               "LPMLV30_CMD_START":
                 IF NOT #statStatesInCurrentMode.resetting AND NOT #statStatesInCurrentMode.idle THEN
                   #StateChangeInProcess := TRUE;
                   #StateRequested := "LPMLV30_STATE_EXECUTE";
                   // Check if valid state for command is in use by current mode
                   IF #statStatesInCurrentMode.starting THEN
                     #statStateInternal := "LPMLV30_STATE_STARTING";
                   ELSE
                     #statStateInternal := "LPMLV30_STATE_EXECUTE";
                   END_IF;
                 ELSE
                   #diagnostics.buffer[#tempDiagnosticsBufferIndexCmd].message := #MSG_CMD_NOT_ALLOWED;
                 END_IF;
               ELSE
                 IF #diagnostics.buffer[#tempDiagnosticsBufferIndexCmd].message = #MSG_NO_MESSAGE THEN // ELSE: Message was already written in head part of message handling
                   #diagnostics.buffer[#tempDiagnosticsBufferIndexCmd].message := #MSG_CMD_NOT_ALLOWED;
                 END_IF;
             END_CASE;
           END_IF;

         "LPMLV30_STATE_UNDEFINED":
           #StateChangeInProcess := FALSE;
           #StateRequested    := "LPMLV30_STATE_STOPPED";
           #statStateInternal := "LPMLV30_STATE_STOPPED";
         ELSE
           ; // Undefined state
       END_CASE;
     END_IF; // End: state machine

     //-------------------------------------------------
     // Message handling for state manager: foot part
     //-------------------------------------------------
     IF #statStateInternal <> #statStateCurrentOld THEN // ELSE: States were not changed
       IF #tempDiagnosticsBufferIndexCmd >= 0 AND #tempDiagnosticsBufferIndexCmd <= "LPMLV30_DIAG_BUFFER_UPPER_LIM" THEN
         IF #diagnostics.buffer[#tempDiagnosticsBufferIndexCmd].message = #MSG_NO_MESSAGE THEN
           #diagnostics.buffer[#tempDiagnosticsBufferIndexCmd].message := #MSG_STATE_CHANGED_SUCCESSFULLY;
         END_IF;
       END_IF;
       IF #tempDiagnosticsBufferIndexSC >= 0 AND #tempDiagnosticsBufferIndexSC <= "LPMLV30_DIAG_BUFFER_UPPER_LIM" THEN
         IF #diagnostics.buffer[#tempDiagnosticsBufferIndexSC].message = #MSG_NO_MESSAGE THEN
           #diagnostics.buffer[#tempDiagnosticsBufferIndexSC].message := #MSG_STATE_CHANGED_SUCCESSFULLY;
         END_IF;
       END_IF;
     END_IF; // End: message handling for state manager: foot part
   END_IF; // End: As from second cycle
   // End: State manager

   //--------------------------------------------------------------------------------------------------
   // Write outputs including boolean interface outputs 
   //--------------------------------------------------------------------------------------------------
   IF #statUnitModeCurrentInternal <> #statUnitModeCurrentInternalOld THEN // Check if new unit mode is selected
     #ProductionModeActive  := FALSE;
     #MaintenanceModeActive := FALSE;
     #ManualModeActive      := FALSE;
     #UserMode01Active      := FALSE;
     #UserMode02Active      := FALSE;
     #UserMode03Active      := FALSE;
     #UserMode04Active      := FALSE;
     #UserMode05Active      := FALSE;
     #UserMode06Active      := FALSE;
     #UserMode07Active      := FALSE;
     #UserMode08Active      := FALSE;
     // #UserMode09Active := FALSE;
     // #UserMode10Active := FALSE;
     // #UserMode11Active := FALSE;
     // #UserMode13Active := FALSE;
     // #UserMode14Active := FALSE;
     // #UserMode15Active := FALSE;
     // #UserMode16Active := FALSE;
     // #UserMode17Active := FALSE;
     // #UserMode18Active := FALSE;
     // #UserMode19Active := FALSE;
     // #UserMode20Active := FALSE;
     // #UserMode21Active := FALSE;
     // #UserMode22Active := FALSE;
     // #UserMode23Active := FALSE;
     // #UserMode24Active := FALSE;
     // #UserMode25Active := FALSE;
     // #UserMode26Active := FALSE;
     // #UserMode27Active := FALSE;
     // #UserMode28Active := FALSE;

     CASE #statUnitModeCurrentInternal OF // Set new bit for current unit mode
       "LPMLV30_MODE_PRODUCTION":
         #ProductionModeActive := TRUE;
       "LPMLV30_MODE_MAINTENANCE":
         #MaintenanceModeActive := TRUE;
       "LPMLV30_MODE_MANUAL":
         #ManualModeActive := TRUE;
       "LPMLV30_MODE_USER_01":
         #UserMode01Active := TRUE;
       "LPMLV30_MODE_USER_02":
         #UserMode02Active := TRUE;
       "LPMLV30_MODE_USER_03":
         #UserMode03Active := TRUE;
       "LPMLV30_MODE_USER_04":
         #UserMode04Active := TRUE;
       "LPMLV30_MODE_USER_05":
         #UserMode05Active := TRUE;
       "LPMLV30_MODE_USER_06":
         #UserMode06Active := TRUE;
       "LPMLV30_MODE_USER_07":
         #UserMode07Active := TRUE;
       "LPMLV30_MODE_USER_08":
         #UserMode08Active := TRUE;
       // LPMLV30_MODE_USER_09:
       //   #UserMode09Active := TRUE;
       // LPMLV30_MODE_USER_10:
       //   #UserMode10Active := TRUE;
       // LPMLV30_MODE_USER_11:
       //   #UserMode11Active := TRUE;
       // LPMLV30_MODE_USER_12:
       //   #UserMode12Active := TRUE;
       // LPMLV30_MODE_USER_13:
       //   #UserMode13Active := TRUE;
       // LPMLV30_MODE_USER_14:
       //   #UserMode14Active := TRUE;
       // LPMLV30_MODE_USER_15:
       //   #UserMode15Active := TRUE;
       // LPMLV30_MODE_USER_16:
       //   #UserMode16Active := TRUE;
       // LPMLV30_MODE_USER_17:
       //   #UserMode17Active := TRUE;
       // LPMLV30_MODE_USER_18:
       //   #UserMode18Active := TRUE;
       // LPMLV30_MODE_USER_19:
       //   #UserMode19Active := TRUE;
       // LPMLV30_MODE_USER_20:
       //   #UserMode20Active := TRUE;
       // LPMLV30_MODE_USER_21:
       //   #UserMode21Active := TRUE;
       // LPMLV30_MODE_USER_22:
       //   #UserMode22Active := TRUE;
       // LPMLV30_MODE_USER_23:
       //   #UserMode23Active := TRUE;
       // LPMLV30_MODE_USER_24:
       //   #UserMode25Active := TRUE;
       // LPMLV30_MODE_USER_25:
       //   #UserMode25Active := TRUE;
       // LPMLV30_MODE_USER_26:
       //   #UserMode26Active := TRUE;
       // LPMLV30_MODE_USER_27:
       //   #UserMode27Active := TRUE;
       // LPMLV30_MODE_USER_28:
       //   #UserMode28Active := TRUE;
       ELSE
         ; // No bit is set
     END_CASE;

     #statUnitModeCurrentInternalOld := #statUnitModeCurrentInternal;
   END_IF;

   IF #statStateInternal <> #statStateInternalOld THEN // Check if new state is selected 
     #StateCurrent := #statStateInternal; // Set output

     // Set states of boolean interface out
     // Delete old state  
     #ClearingStateActive     := FALSE;
     #StoppedStateActive      := FALSE;
     #StartingStateActive     := FALSE;
     #IdleStateActive         := FALSE;
     #SuspendedStateActive    := FALSE;
     #ExecuteStateActive      := FALSE;
     #StoppingStateActive     := FALSE;
     #AbortingStateActive     := FALSE;
     #AbortedStateActive      := FALSE;
     #HoldingStateActive      := FALSE;
     #HeldStateActive         := FALSE;
     #UnholdingStateActive    := FALSE;
     #SuspendingStateActive   := FALSE;
     #UnsuspendingStateActive := FALSE;
     #ResettingStateActive    := FALSE;
     #CompletingStateActive   := FALSE;
     #CompleteStateActive     := FALSE;

     // Set new state
     CASE #statStateInternal OF
       "LPMLV30_STATE_CLEARING":
         #ClearingStateActive := TRUE;
       "LPMLV30_STATE_STOPPED":
         #StoppedStateActive := TRUE;
       "LPMLV30_STATE_STARTING":
         #StartingStateActive := TRUE;
       "LPMLV30_STATE_IDLE":
         #IdleStateActive := TRUE;
       "LPMLV30_STATE_SUSPENDED":
         #SuspendedStateActive := TRUE;
       "LPMLV30_STATE_EXECUTE":
         #ExecuteStateActive := TRUE;
       "LPMLV30_STATE_STOPPING":
         #StoppingStateActive := TRUE;
       "LPMLV30_STATE_ABORTING":
         #AbortingStateActive := TRUE;
       "LPMLV30_STATE_ABORTED":
         #AbortedStateActive := TRUE;
       "LPMLV30_STATE_HOLDING":
         #HoldingStateActive := TRUE;
       "LPMLV30_STATE_HELD":
         #HeldStateActive := TRUE;
       "LPMLV30_STATE_UNHOLDING":
         #UnholdingStateActive := TRUE;
       "LPMLV30_STATE_SUSPENDING":
         #SuspendingStateActive := TRUE;
       "LPMLV30_STATE_UNSUSPENDING":
         #UnsuspendingStateActive := TRUE;
       "LPMLV30_STATE_RESETTING":
         #ResettingStateActive := TRUE;
       "LPMLV30_STATE_COMPLETING":
         #CompletingStateActive := TRUE;
       "LPMLV30_STATE_COMPLETE":
         #CompleteStateActive := TRUE;
       ELSE
         ;
     END_CASE; // End: Set new state

     #statStateInternalOld := #statStateInternal;
   END_IF;// End: Write boolean interface outputs

   #diagnostics.bufferIndex := #tempDiagnosticsBufferIndex; // Temporary variable is used during block execution -> Copy back/Set output
   IF #statFirstCycle THEN
     #statFirstCycle := FALSE;
   END_IF;

   // Save values for edge detection
   IF #statUnitModeChangeRequest THEN
     #statUnitModeOld := #statUnitMode;
   END_IF;
   IF #statCmdChangeRequest THEN
     #statCntrlCmdOld := #tempCntrlCmd;
   END_IF;
   IF #statStateInternal <> #statStateCurrentOld THEN
     #statStateCurrentOld := #statStateInternal;
   END_IF;

   //============================================================================================================
   // End of function block: LPMLV30_UnitModeStateManager
   //============================================================================================================
END_FUNCTION_BLOCK

FUNCTION_BLOCK "LPMLV30_UnitModeStateTimes"   // FB30101, SCL
TITLE = LPMLV30_UnitModeStateTimes
{ S7_Optimized_Access := 'TRUE' }
AUTHOR : APC_ERLF
FAMILY : OMAC
// Support: tech.team.motioncontrol@siemens.com 
// Fax: +49 (0) 9131/98-1297
   VAR_INPUT
      UnitModeCurrent : DInt := 0;   // Current unit mode
      StateCurrent : DInt := 0;   // Current state
      resetTimes : Bool := false;   // State change from FALSE to TRUE (rising edge) resets unit mode/state times and cumulative times
   END_VAR
   VAR_OUTPUT
      ModeCurrentTime : Array[0.."LPMLV30_MODES_UPPER_LIM"] of DInt;   // Current time for all modes in seconds
      ModeCumulativeTime : Array[0.."LPMLV30_MODES_UPPER_LIM"] of DInt;   // Cumulative time for all modes in seconds
      StateCurrentTime : Array[0.."LPMLV30_MODES_UPPER_LIM", 0.."LPMLV30_STATES_UPPER_LIM"] of DInt;   // Current time for all states in seconds
      StateCumulativeTime : Array[0.."LPMLV30_MODES_UPPER_LIM", 0.."LPMLV30_STATES_UPPER_LIM"] of DInt;   // Cumulative time for all states in seconds
      actualTimeCurrentMode : DInt;   // Actual time for current mode in seconds
      cumulativeTimeCurrentMode : DInt;   // Cumulative time for current mode in seconds
      actualTimeCurrentStates : Array[0.."LPMLV30_STATES_UPPER_LIM"] of DInt;   // Actual time for all states in current mode in seconds
      cumulativeTimeCurrentStates : Array[0.."LPMLV30_STATES_UPPER_LIM"] of DInt;   // Cumulative time for all states in current mode in seconds
      AccTimeSinceReset : DInt;   // Accumulated time since last reset in seconds
   END_VAR
   VAR
      statUnitModeCurrentOld : DInt := 0;   // For edge detection
      statStateCurrentOld : DInt := 0;   // For edge detection
      statResetTimesOld : Bool := false;   // For edge detection
      statStartingPointMeasureRuntime : LReal := 0.0;   // Saved value of runtime system function
      statRuntime : LReal := 0.0;   // Runtime variable
      statFirstCycle : Bool := true;   // First cycle of run
   END_VAR
   VAR_TEMP
      tempI : Int;   // Loop counter
      tempJ : Int;   // Loop counter
      tempMeasuredRuntime : LReal;   // Return value of RUNTIME instruction
      tempRuntimeIntegerPart : DInt;   // Runtime variable (integer part)
      tempUnitModeCurrent : DInt;   // Verified input value
      tempStateCurrent : DInt;   // Verified input value
   END_VAR
BEGIN
   //============================================================================================================
   // SIEMENS AG
   // (c)Copyright 2015 All Rights Reserved
   //------------------------------------------------------------------------------------------------------------
   // Library: LPMLV30
   // Tested with: S7-1200 with FW version V4.1, S7-1500 with FW version V1.7
   // Engineering: TIA Portal V13 SP1
   // Restrictions: ---
   // Requirements: S7-1200 / S7-1500
   // Functionality: Determination of unit modes and states times (current and also cumulative times)
   //------------------------------------------------------------------------------------------------------------
   // Change log table:
   // Version  Date        Expert in charge    Changes applied
   // 03.00.01 29.05.2015  RK                  First released version 
   //============================================================================================================
   // Function block: LPMLV30_UnitModeStateTimes
   //============================================================================================================

   IF #statFirstCycle OR (#resetTimes AND NOT #statResetTimesOld) THEN
     // Reset times structures
     FOR #tempI := "LPMLV30_MODE_INVALID" TO "LPMLV30_MODES_UPPER_LIM" DO
       #ModeCurrentTime[#tempI] := 0;
       IF NOT #statFirstCycle THEN // Do only with rising edge at resetTimes
         #ModeCumulativeTime[#tempI] := 0;
       END_IF;
       FOR #tempJ := "LPMLV30_STATE_UNDEFINED" TO "LPMLV30_STATES_UPPER_LIM" DO
         #StateCurrentTime[#tempI, #tempJ] := 0;
         IF NOT #statFirstCycle THEN // Do only with rising edge at resetTimes
           #StateCumulativeTime[#tempI, #tempJ] := 0;
         END_IF;
       END_FOR;
     END_FOR;
     IF NOT #statFirstCycle THEN // Do only with rising edge at resetTimes
       #AccTimeSinceReset := 0;
     END_IF;

     // Reset additional outputs
     #actualTimeCurrentMode := 0;
     IF NOT #statFirstCycle THEN // Do only with rising edge at resetTimes
       #cumulativeTimeCurrentMode := 0;
     END_IF;
     FOR #tempI := "LPMLV30_STATE_UNDEFINED" TO "LPMLV30_STATES_UPPER_LIM" DO
       #actualTimeCurrentStates[#tempI] := 0;
       IF NOT #statFirstCycle THEN // Do only with rising edge at resetTimes
         #cumulativeTimeCurrentStates[#tempI] := 0;
       END_IF;
     END_FOR;

     // Set starting point for calculation of elapsed seconds
     #tempMeasuredRuntime := RUNTIME(#statStartingPointMeasureRuntime);
     #statRuntime := 0.0;

     IF #statFirstCycle THEN
       #statFirstCycle := FALSE;
       RETURN; // Nothing else in this cycle to avoid runtime peaks
     END_IF;
   END_IF;

   // Inputs UnitModeCurrent and StateCurrent
   #tempUnitModeCurrent := #UnitModeCurrent;
   #tempStateCurrent    := #StateCurrent;

   // Measure program runtime
   #tempMeasuredRuntime := RUNTIME(#statStartingPointMeasureRuntime);
   IF #tempMeasuredRuntime > 0.0 THEN //value OK
     #statRuntime := #statRuntime + #tempMeasuredRuntime;
   END_IF;

   // Check if at least one second has been reached
   IF #statRuntime > 1.0 THEN
     #tempRuntimeIntegerPart := TRUNC_DINT(#statRuntime);

     IF #statUnitModeCurrentOld >= "LPMLV30_MODE_INVALID" AND #statUnitModeCurrentOld <= "LPMLV30_MODES_UPPER_LIM" THEN
       //DINT overflow is not taken into account, because DINT in seconds means approx. 68 years
       #ModeCurrentTime[#statUnitModeCurrentOld]    := #ModeCurrentTime[#statUnitModeCurrentOld]    + #tempRuntimeIntegerPart;
       #ModeCumulativeTime[#statUnitModeCurrentOld] := #ModeCumulativeTime[#statUnitModeCurrentOld] + #tempRuntimeIntegerPart;

       IF #statStateCurrentOld >= "LPMLV30_STATE_UNDEFINED" AND #statStateCurrentOld <= "LPMLV30_STATES_UPPER_LIM" THEN
         //DINT overflow is not taken into account, because DINT in seconds means approx. 68 years
         #StateCurrentTime[#statUnitModeCurrentOld, #statStateCurrentOld]    := #StateCurrentTime[#statUnitModeCurrentOld, #statStateCurrentOld]    + #tempRuntimeIntegerPart;
         #StateCumulativeTime[#statUnitModeCurrentOld, #statStateCurrentOld] := #StateCumulativeTime[#statUnitModeCurrentOld, #statStateCurrentOld] + #tempRuntimeIntegerPart;
       END_IF;
     END_IF;

     //DINT overflow is not taken into account, because DINT in seconds means approx. 68 years
     #AccTimeSinceReset := #AccTimeSinceReset + #tempRuntimeIntegerPart;

     #statRuntime := #statRuntime - #tempRuntimeIntegerPart; //fractional part of runtime variable for next cycle
   END_IF;

   // Check if new unitMode is selected
   IF #tempUnitModeCurrent <> #statUnitModeCurrentOld THEN
     IF #tempUnitModeCurrent >= "LPMLV30_MODE_INVALID" AND #tempUnitModeCurrent <= "LPMLV30_MODES_UPPER_LIM" THEN
       #ModeCurrentTime[#tempUnitModeCurrent] := 0;
       IF #tempStateCurrent >= "LPMLV30_STATE_UNDEFINED" AND #tempStateCurrent <= "LPMLV30_STATES_UPPER_LIM" THEN
         #StateCurrentTime[#tempUnitModeCurrent, #tempStateCurrent] := 0;
       END_IF;
     END_IF;

   // Check if new state is selected   
   ELSIF #tempStateCurrent <> #statStateCurrentOld THEN
     IF #tempUnitModeCurrent >= "LPMLV30_MODE_INVALID"    AND #tempUnitModeCurrent <= "LPMLV30_MODES_UPPER_LIM" AND
        #tempStateCurrent    >= "LPMLV30_STATE_UNDEFINED" AND #tempStateCurrent    <= "LPMLV30_STATES_UPPER_LIM"
     THEN
       #StateCurrentTime[#tempUnitModeCurrent, #tempStateCurrent] := 0;
     END_IF;
   END_IF;

   // Update additional outputs
   IF #tempUnitModeCurrent >= "LPMLV30_MODE_INVALID" AND #tempUnitModeCurrent <= "LPMLV30_MODES_UPPER_LIM" THEN
     #actualTimeCurrentMode     := #ModeCurrentTime[#tempUnitModeCurrent];
     #cumulativeTimeCurrentMode := #ModeCumulativeTime[#tempUnitModeCurrent];
     IF #tempStateCurrent >= "LPMLV30_STATE_UNDEFINED" AND #tempStateCurrent <= "LPMLV30_STATES_UPPER_LIM" THEN
       #actualTimeCurrentStates     := #StateCurrentTime[#tempUnitModeCurrent];
       #cumulativeTimeCurrentStates := #StateCumulativeTime[#tempUnitModeCurrent];
     ELSE
       FOR #tempI := "LPMLV30_STATE_UNDEFINED" TO "LPMLV30_STATES_UPPER_LIM" DO
         #actualTimeCurrentStates[#tempI] := 0;
         #cumulativeTimeCurrentStates[#tempI] := 0;
       END_FOR;
     END_IF;
   ELSE
     #actualTimeCurrentMode     := 0;
     #cumulativeTimeCurrentMode := 0;

     FOR #tempI := "LPMLV30_STATE_UNDEFINED" TO "LPMLV30_STATES_UPPER_LIM" DO
       #actualTimeCurrentStates[#tempI]     := 0;
       #cumulativeTimeCurrentStates[#tempI] := 0;
     END_FOR;
   END_IF;

   // Save values for state change detection
   #statResetTimesOld      := #resetTimes;
   #statUnitModeCurrentOld := #tempUnitModeCurrent;
   #statStateCurrentOld    := #tempStateCurrent;

   //============================================================================================================
   // End of Function block: LPMLV30_UnitModeStateTimes
   //============================================================================================================
END_FUNCTION_BLOCK

FUNCTION "LPMLV30_ConfigureDisabledUnitModes" : Void   // FC30100, SCL
TITLE = LPMLV30_ConfigureDisabledUnitModes
{ S7_Optimized_Access := 'TRUE' }
AUTHOR : APC_ERLF
FAMILY : OMAC
// Support: tech.team.motioncontrol@siemens.com 
// Fax: +49 (0) 9131/98-1297
   VAR_INPUT
      ProductionModeDisable : Bool;   // TRUE: Disable unit mode Production
      MaintenanceModeDisable : Bool;   // TRUE: Disable unit mode Maintenance
      UserMode01Disable : Bool;   // TRUE: Disable user-defined unit mode 01
      UserMode02Disable : Bool;   // TRUE: Disable user-defined unit mode 02
      UserMode03Disable : Bool;   // TRUE: Disable user-defined unit mode 03
      UserMode04Disable : Bool;   // TRUE: Disable user-defined unit mode 04
      UserMode05Disable : Bool;   // TRUE: Disable user-defined unit mode 05
      UserMode06Disable : Bool;   // TRUE: Disable user-defined unit mode 06
      UserMode07Disable : Bool;   // TRUE: Disable user-defined unit mode 07
      UserMode08Disable : Bool;   // TRUE: Disable user-defined unit mode 08
   END_VAR
   VAR_OUTPUT
      disabledUnitModes : Array[0.."LPMLV30_MAX_MODES_UPPER_LIM"] of Bool;   // Disabled unit modes configuration
   END_VAR
   VAR_TEMP
      tempI : Int;   // Temporary Index
   END_VAR
   // Ret_Val : Function without return value
BEGIN
   //============================================================================================================
   // SIEMENS AG
   // (c)Copyright 2015 All Rights Reserved
   //------------------------------------------------------------------------------------------------------------
   // Library: LPMLV30
   // Tested with: S7-1200 with FW version V4.1, S7-1500 with FW version V1.7
   // Engineering: TIA Portal V13 SP1
   // Restrictions: ---
   // Requirements: S7-1200 / S7-1500
   // Functionality: The function generates the unit mode configuration as Array[] of Bool.
   //------------------------------------------------------------------------------------------------------------
   // Change log table:
   // Version  Date        Expert in charge    Changes applied
   // 03.00.01 29.05.2015  RK                  First released version 
   //============================================================================================================
   // Function: LPMLV30_ConfigureDisabledUnitModes
   //============================================================================================================

   // Initialize unitMode configuration
   FOR #tempI := 0 TO "LPMLV30_MAX_MODES_UPPER_LIM" DO
     #disabledUnitModes[#tempI] := TRUE;
   END_FOR;

   // Set unitMode configuration
   #disabledUnitModes["LPMLV30_MODE_INVALID"]     := FALSE;
   #disabledUnitModes["LPMLV30_MODE_PRODUCTION"]  := #ProductionModeDisable;
   #disabledUnitModes["LPMLV30_MODE_MAINTENANCE"] := #MaintenanceModeDisable;
   #disabledUnitModes["LPMLV30_MODE_MANUAL"]      := FALSE;
   #disabledUnitModes["LPMLV30_MODE_USER_01"]     := #UserMode01Disable;
   #disabledUnitModes["LPMLV30_MODE_USER_02"]     := #UserMode02Disable;
   #disabledUnitModes["LPMLV30_MODE_USER_03"]     := #UserMode03Disable;
   #disabledUnitModes["LPMLV30_MODE_USER_04"]     := #UserMode04Disable;
   #disabledUnitModes["LPMLV30_MODE_USER_05"]     := #UserMode05Disable;
   #disabledUnitModes["LPMLV30_MODE_USER_06"]     := #UserMode06Disable;
   #disabledUnitModes["LPMLV30_MODE_USER_07"]     := #UserMode07Disable;
   #disabledUnitModes["LPMLV30_MODE_USER_08"]     := #UserMode08Disable;

   //============================================================================================================
   // End of function: LPMLV30_ConfigureDisabledUnitModes
   //============================================================================================================
END_FUNCTION

FUNCTION "LPMLV30_ConfigureDisabledStates" : Void   // FC30101, SCL
TITLE = LPMLV30_ConfigureDisabledStates
{ S7_Optimized_Access := 'TRUE' }
AUTHOR : APC_ERLF
FAMILY : OMAC
// Support: tech.team.motioncontrol@siemens.com 
// Fax: +49 (0) 9131/98-1297
   VAR_INPUT
      HoldingDisable : Bool;   // TRUE: Disable state Holding
      HeldDisable : Bool;   // TRUE: Disable state Held
      UnholdingDisable : Bool;   // TRUE: Disable state Unholding
      SuspendingDisable : Bool;   // TRUE: Disable state Suspending
      SuspendedDisable : Bool;   // TRUE: Disable state Suspended
      UnsuspendingDisable : Bool;   // TRUE: Disable state Unsuspending
      CompletingDisable : Bool;   // TRUE: Disable state Completing
      CompleteDisable : Bool;   // TRUE: Disable state Complete
   END_VAR
   VAR_OUTPUT
      disabledStates : DInt;   // Disabled states configuration for one unit mode
   END_VAR
   // Ret_Val : Function without return value
   VAR CONSTANT
      DISABLE_ALL_STATES : DWord := 16#FFFF_FFFF;   // Disable all states
   END_VAR
BEGIN
   //============================================================================================================
   // SIEMENS AG
   // (c)Copyright 2015 All Rights Reserved
   //------------------------------------------------------------------------------------------------------------
   // Library: LPMLV30
   // Tested with: S7-1200 with FW version V4.1, S7-1500 with FW version V1.7
   // Engineering: TIA Portal V13 SP1
   // Restrictions: ---
   // Requirements: S7-1200 / S7-1500
   // Functionality: The function generates a double integer value which represents the state configuration
   //                for one unit mode.
   //------------------------------------------------------------------------------------------------------------
   // Change log table:
   // Version  Date        Expert in charge    Changes applied
   // 03.00.01 29.05.2015  RK                  First released version 
   //============================================================================================================
   // Function: LPMLV30_ConfigureDisabledStates
   //============================================================================================================

   #disabledStates := DWORD_TO_DINT(#DISABLE_ALL_STATES);

   #disabledStates.%X0  := FALSE; // Undefined state is mandatory
   #disabledStates.%X1  := FALSE; // Clearing state is mandatory
   #disabledStates.%X2  := FALSE; // Stopped state is mandatory
   #disabledStates.%X3  := FALSE; // Starting state is mandatory
   #disabledStates.%X4  := FALSE; // Idle state is mandatory
   #disabledStates.%X5  := #SuspendedDisable;
   #disabledStates.%X6  := FALSE; // Execute state is mandatory
   #disabledStates.%X7  := FALSE; // Stopping state is mandatory
   #disabledStates.%X8  := FALSE; // Aborting state is mandatory
   #disabledStates.%X9  := FALSE; // Aborted state is mandatory
   #disabledStates.%X10 := #HoldingDisable;
   #disabledStates.%X11 := #HeldDisable;
   #disabledStates.%X12 := #UnholdingDisable;
   #disabledStates.%X13 := #SuspendingDisable;
   #disabledStates.%X14 := #UnsuspendingDisable;
   #disabledStates.%X15 := FALSE; // Resetting state is mandatory
   #disabledStates.%X16 := #CompletingDisable;
   #disabledStates.%X17 := #CompleteDisable;

   //============================================================================================================
   // End of function: LPMLV30_ConfigureDisabledStates
   //============================================================================================================
END_FUNCTION

FUNCTION "LPMLV30_GetUnitModeStateNamesAsString" : Void   // FC30102, SCL
TITLE = LPMLV30_GetUnitModeStateNamesAsString
{ S7_Optimized_Access := 'TRUE' }
AUTHOR : APC_ERLF
FAMILY : OMAC
// Support: tech.team.motioncontrol@siemens.com 
// Fax: +49 (0) 9131/98-1297
   VAR_INPUT
      UnitModeCurrent : DInt;   // Current unit mode
      StateCurrent : DInt;   // Current state
      language : Int;   // Requested language (LPMLV30_LANGUAGE_1, LPMLV30_LANGUAGE_2, ...)
      namesConfiguration : "typeLPMLV30_NamesConfiguration";   // All names of unit modes and states (in different languages)
   END_VAR
   VAR_OUTPUT
      unitModeCurrentName : String;   // Name of current unit mode in the requested language
      stateCurrentName : String;   // Name of current state in the requested language
   END_VAR
   VAR_TEMP
      tempUnitModeCurrent : DInt;   // Current unit mode
      tempStateCurrent : DInt;   // Current state
      tempLanguage : Int;   // Requested language
   END_VAR
   // Ret_Val : Function without return value
BEGIN
   //============================================================================================================
   // SIEMENS AG
   // (c)Copyright 2015 All Rights Reserved
   //------------------------------------------------------------------------------------------------------------
   // Library: LPMLV30
   // Tested with: S7-1200 with FW version V4.1, S7-1500 with FW version V1.7
   // Engineering: TIA Portal V13 SP1
   // Restrictions: ---
   // Requirements: S7-1200 / S7-1500
   // Functionality: Gets the names for current unit mode and state in one language 
   //                corresponding to the names configuration
   //------------------------------------------------------------------------------------------------------------
   // Change log table:
   // Version  Date        Expert in charge    Changes applied
   // 03.00.01 29.05.2015  RK                  First released version 
   //============================================================================================================
   // Function: LPMLV30_GetUnitModeStateNamesAsString
   //============================================================================================================

   #tempUnitModeCurrent := #UnitModeCurrent;
   #tempStateCurrent    := #StateCurrent;
   #tempLanguage        := #language;

   IF #tempUnitModeCurrent < 0 OR #tempUnitModeCurrent > "LPMLV30_MODES_UPPER_LIM" THEN
     #tempUnitModeCurrent := "LPMLV30_MODE_INVALID";
   END_IF;
   IF #tempStateCurrent < 0 OR #tempStateCurrent > "LPMLV30_STATES_UPPER_LIM" THEN
     #tempStateCurrent := "LPMLV30_STATE_UNDEFINED";
   END_IF;
   IF #tempLanguage < 0 OR #tempLanguage > "LPMLV30_LANGUAGES_UPPER_LIM" THEN
     #tempLanguage := "LPMLV30_LANGUAGE_1";
   END_IF;

   #unitModeCurrentName := #namesConfiguration.unitModesNames[#tempLanguage, #tempUnitModeCurrent];
   #stateCurrentName    := #namesConfiguration.statesNames[#tempLanguage, #tempStateCurrent];

   //============================================================================================================
   // End of function: LPMLV30_GetUnitModeStateNamesAsString
   //============================================================================================================
END_FUNCTION

// folder: _UN01_Palletizer

FUNCTION_BLOCK "UN_00_Main"   // FB31620, LAD
TITLE = UN_00_Main
{ S7_Optimized_Access := 'TRUE' }
AUTHOR : tech.team.motioncontrol@siemens.com
FAMILY : CPG
VERSION : 1.0
// Support: tech.team.motioncontrol@siemens.com
// Fax: +49 (0) 9131/98-1297
   VAR
      instPackML_ModuleSum : "UN_01_PackML_ModuleSum";   // PackML Module Summation Logic of EM-level command and state complete's to unit level
      instPackML : "UN_02_PackML";
      instLineComm : "UN_03_LineComm";
      instEventControl : "UN_04_EventControl";
      instEventSummation : "UN_05_EventSummation";
      instMiscFunctions : "UN_06_MiscFunctions";
      instRecipeControl : "UN_07_RecipeControl";
   END_VAR
   VAR_TEMP   // added for the SCL form of the ladder/FBD networks
      _w1 : Bool;
   END_VAR
BEGIN

REGION Network 1: Call the PackML Module Summation Logic
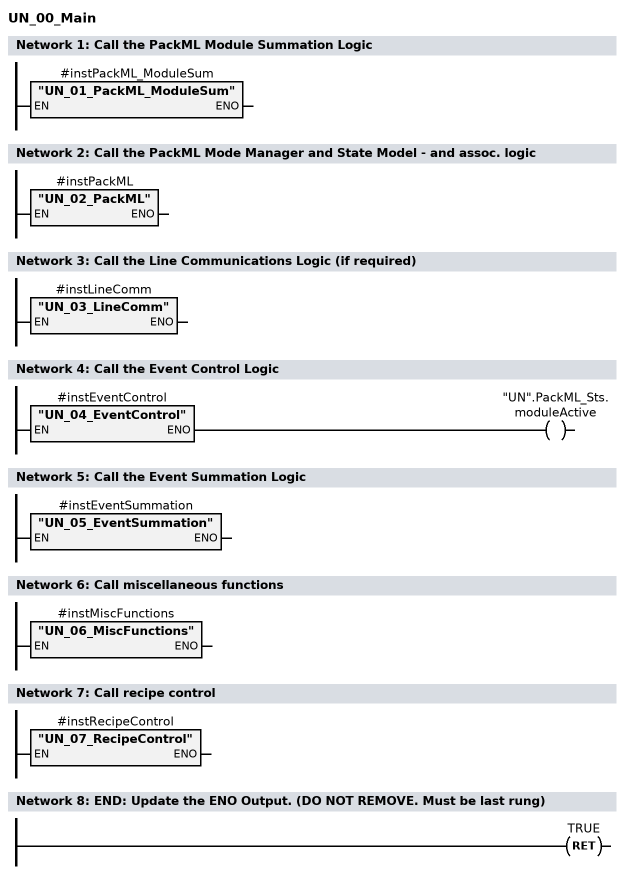
   RUNG wire#powerrail
      #instPackML_ModuleSum()
   END_RUNG
   // the same network as SCL:
   #instPackML_ModuleSum();   // "UN_01_PackML_ModuleSum"
END_REGION

REGION Network 2: Call the PackML Mode Manager and State Model - and assoc. logic
   RUNG wire#powerrail
      #instPackML()
   END_RUNG
   // the same network as SCL:
   #instPackML();   // "UN_02_PackML"
END_REGION

REGION Network 3: Call the Line Communications Logic (if required)
   RUNG wire#powerrail
      #instLineComm()
   END_RUNG
   // the same network as SCL:
   #instLineComm();   // "UN_03_LineComm"
END_REGION

REGION Network 4: Call the Event Control Logic
   RUNG wire#powerrail
      #instEventControl()
      Coil( "UN".PackML_Sts.moduleActive )
   END_RUNG
   // the same network as SCL:
   #instEventControl(ENO => #_w1);   // "UN_04_EventControl"
   "UN".PackML_Sts.moduleActive := #_w1;
END_REGION

REGION Network 5: Call the Event Summation Logic
   RUNG wire#powerrail
      #instEventSummation()
   END_RUNG
   // the same network as SCL:
   #instEventSummation();   // "UN_05_EventSummation"
END_REGION

REGION Network 6: Call miscellaneous functions
   RUNG wire#powerrail
      #instMiscFunctions()
   END_RUNG
   // the same network as SCL:
   #instMiscFunctions();   // "UN_06_MiscFunctions"
END_REGION

REGION Network 7: Call recipe control
   RUNG wire#powerrail
      #instRecipeControl()
   END_RUNG
   // the same network as SCL:
   #instRecipeControl();   // "UN_07_RecipeControl"
END_REGION

REGION Network 8: END: Update the ENO Output. (DO NOT REMOVE. Must be last rung)
   RUNG wire#powerrail
      ReturnCoil( TRUE )
   END_RUNG
   // the same network as SCL:
   ENO := TRUE;
   RETURN;
END_REGION
END_FUNCTION_BLOCK

FUNCTION_BLOCK "UN_01_PackML_ModuleSum"   // FB31621, LAD
TITLE = UN_01_PackML_ModuleSummation
{ S7_Optimized_Access := 'TRUE' }
AUTHOR : tech.team.motioncontrol@siemens.com
FAMILY : CPG
VERSION : 1.0
// Support: tech.team.motioncontrol@siemens.com
// Fax: +49 (0) 9131/98-1297
   VAR
      statDummyBool : Bool;   // dummy bool - placeholder
   END_VAR
BEGIN

REGION Network 1: UN - Reset Command
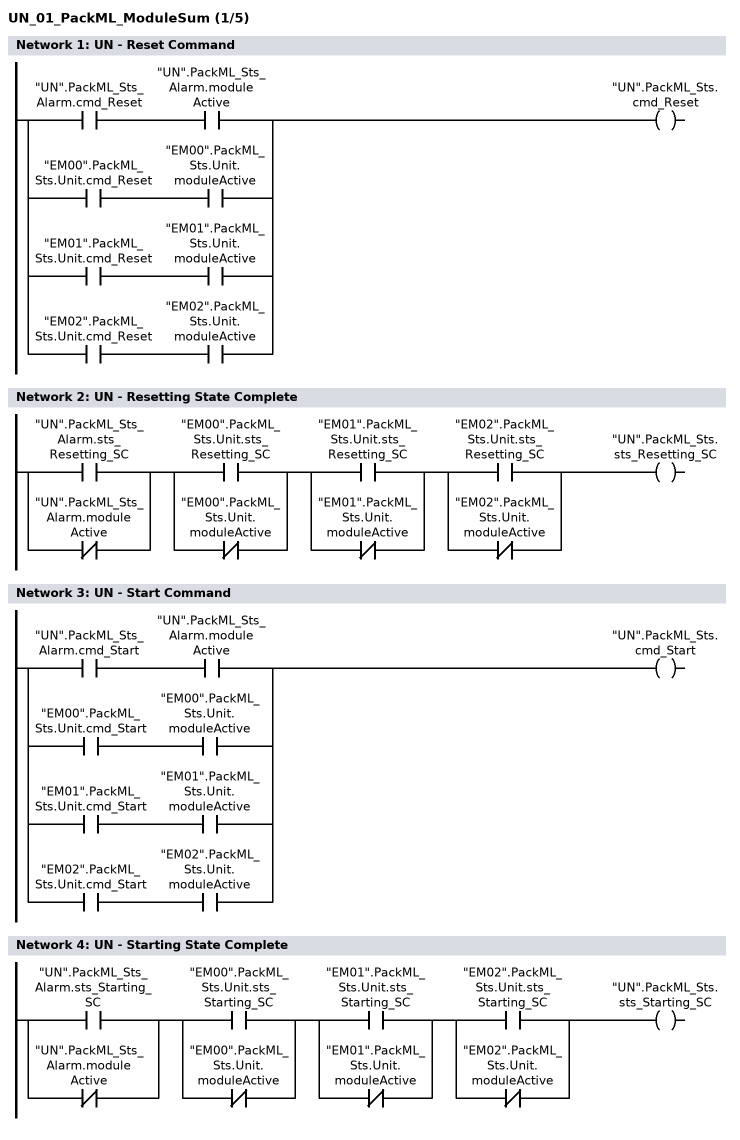
   RUNG wire#powerrail
      Contact( "UN".PackML_Sts_Alarm.cmd_Reset )
      Contact( "UN".PackML_Sts_Alarm.moduleActive )
      wire#w1
      Coil( "UN".PackML_Sts.cmd_Reset )
   END_RUNG
   RUNG wire#powerrail
      Contact( "EM00".PackML_Sts.Unit.cmd_Reset )
      Contact( "EM00".PackML_Sts.Unit.moduleActive )
   END_RUNG wire#w1
   RUNG wire#powerrail
      Contact( "EM01".PackML_Sts.Unit.cmd_Reset )
      Contact( "EM01".PackML_Sts.Unit.moduleActive )
   END_RUNG wire#w1
   RUNG wire#powerrail
      Contact( "EM02".PackML_Sts.Unit.cmd_Reset )
      Contact( "EM02".PackML_Sts.Unit.moduleActive )
   END_RUNG wire#w1
   // the same network as SCL:
   "UN".PackML_Sts.cmd_Reset := ("UN".PackML_Sts_Alarm.cmd_Reset AND "UN".PackML_Sts_Alarm.moduleActive) OR ("EM00".PackML_Sts.Unit.cmd_Reset AND "EM00".PackML_Sts.Unit.moduleActive) OR ("EM01".PackML_Sts.Unit.cmd_Reset AND "EM01".PackML_Sts.Unit.moduleActive) OR ("EM02".PackML_Sts.Unit.cmd_Reset AND "EM02".PackML_Sts.Unit.moduleActive);
END_REGION

REGION Network 2: UN - Resetting State Complete
   RUNG wire#powerrail
      Contact( "UN".PackML_Sts_Alarm.sts_Resetting_SC )
      wire#w1
      Contact( "EM00".PackML_Sts.Unit.sts_Resetting_SC )
      wire#w2
      Contact( "EM01".PackML_Sts.Unit.sts_Resetting_SC )
      wire#w3
      Contact( "EM02".PackML_Sts.Unit.sts_Resetting_SC )
      wire#w4
      Coil( "UN".PackML_Sts.sts_Resetting_SC )
   END_RUNG
   RUNG wire#powerrail
      I_Contact( "UN".PackML_Sts_Alarm.moduleActive )
   END_RUNG wire#w1
   RUNG wire#w1
      I_Contact( "EM00".PackML_Sts.Unit.moduleActive )
   END_RUNG wire#w2
   RUNG wire#w2
      I_Contact( "EM01".PackML_Sts.Unit.moduleActive )
   END_RUNG wire#w3
   RUNG wire#w3
      I_Contact( "EM02".PackML_Sts.Unit.moduleActive )
   END_RUNG wire#w4
   // the same network as SCL:
   "UN".PackML_Sts.sts_Resetting_SC := ("UN".PackML_Sts_Alarm.sts_Resetting_SC OR NOT "UN".PackML_Sts_Alarm.moduleActive) AND ("EM00".PackML_Sts.Unit.sts_Resetting_SC OR NOT "EM00".PackML_Sts.Unit.moduleActive) AND ("EM01".PackML_Sts.Unit.sts_Resetting_SC OR NOT "EM01".PackML_Sts.Unit.moduleActive) AND ("EM02".PackML_Sts.Unit.sts_Resetting_SC OR NOT "EM02".PackML_Sts.Unit.moduleActive);
END_REGION

REGION Network 3: UN - Start Command
   RUNG wire#powerrail
      Contact( "UN".PackML_Sts_Alarm.cmd_Start )
      Contact( "UN".PackML_Sts_Alarm.moduleActive )
      wire#w1
      Coil( "UN".PackML_Sts.cmd_Start )
   END_RUNG
   RUNG wire#powerrail
      Contact( "EM00".PackML_Sts.Unit.cmd_Start )
      Contact( "EM00".PackML_Sts.Unit.moduleActive )
   END_RUNG wire#w1
   RUNG wire#powerrail
      Contact( "EM01".PackML_Sts.Unit.cmd_Start )
      Contact( "EM01".PackML_Sts.Unit.moduleActive )
   END_RUNG wire#w1
   RUNG wire#powerrail
      Contact( "EM02".PackML_Sts.Unit.cmd_Start )
      Contact( "EM02".PackML_Sts.Unit.moduleActive )
   END_RUNG wire#w1
   // the same network as SCL:
   "UN".PackML_Sts.cmd_Start := ("UN".PackML_Sts_Alarm.cmd_Start AND "UN".PackML_Sts_Alarm.moduleActive) OR ("EM00".PackML_Sts.Unit.cmd_Start AND "EM00".PackML_Sts.Unit.moduleActive) OR ("EM01".PackML_Sts.Unit.cmd_Start AND "EM01".PackML_Sts.Unit.moduleActive) OR ("EM02".PackML_Sts.Unit.cmd_Start AND "EM02".PackML_Sts.Unit.moduleActive);
END_REGION

REGION Network 4: UN - Starting State Complete
   RUNG wire#powerrail
      Contact( "UN".PackML_Sts_Alarm.sts_Starting_SC )
      wire#w1
      Contact( "EM00".PackML_Sts.Unit.sts_Starting_SC )
      wire#w2
      Contact( "EM01".PackML_Sts.Unit.sts_Starting_SC )
      wire#w3
      Contact( "EM02".PackML_Sts.Unit.sts_Starting_SC )
      wire#w4
      Coil( "UN".PackML_Sts.sts_Starting_SC )
   END_RUNG
   RUNG wire#powerrail
      I_Contact( "UN".PackML_Sts_Alarm.moduleActive )
   END_RUNG wire#w1
   RUNG wire#w1
      I_Contact( "EM00".PackML_Sts.Unit.moduleActive )
   END_RUNG wire#w2
   RUNG wire#w2
      I_Contact( "EM01".PackML_Sts.Unit.moduleActive )
   END_RUNG wire#w3
   RUNG wire#w3
      I_Contact( "EM02".PackML_Sts.Unit.moduleActive )
   END_RUNG wire#w4
   // the same network as SCL:
   "UN".PackML_Sts.sts_Starting_SC := ("UN".PackML_Sts_Alarm.sts_Starting_SC OR NOT "UN".PackML_Sts_Alarm.moduleActive) AND ("EM00".PackML_Sts.Unit.sts_Starting_SC OR NOT "EM00".PackML_Sts.Unit.moduleActive) AND ("EM01".PackML_Sts.Unit.sts_Starting_SC OR NOT "EM01".PackML_Sts.Unit.moduleActive) AND ("EM02".PackML_Sts.Unit.sts_Starting_SC OR NOT "EM02".PackML_Sts.Unit.moduleActive);
END_REGION

REGION Network 5: UN - Stop Command
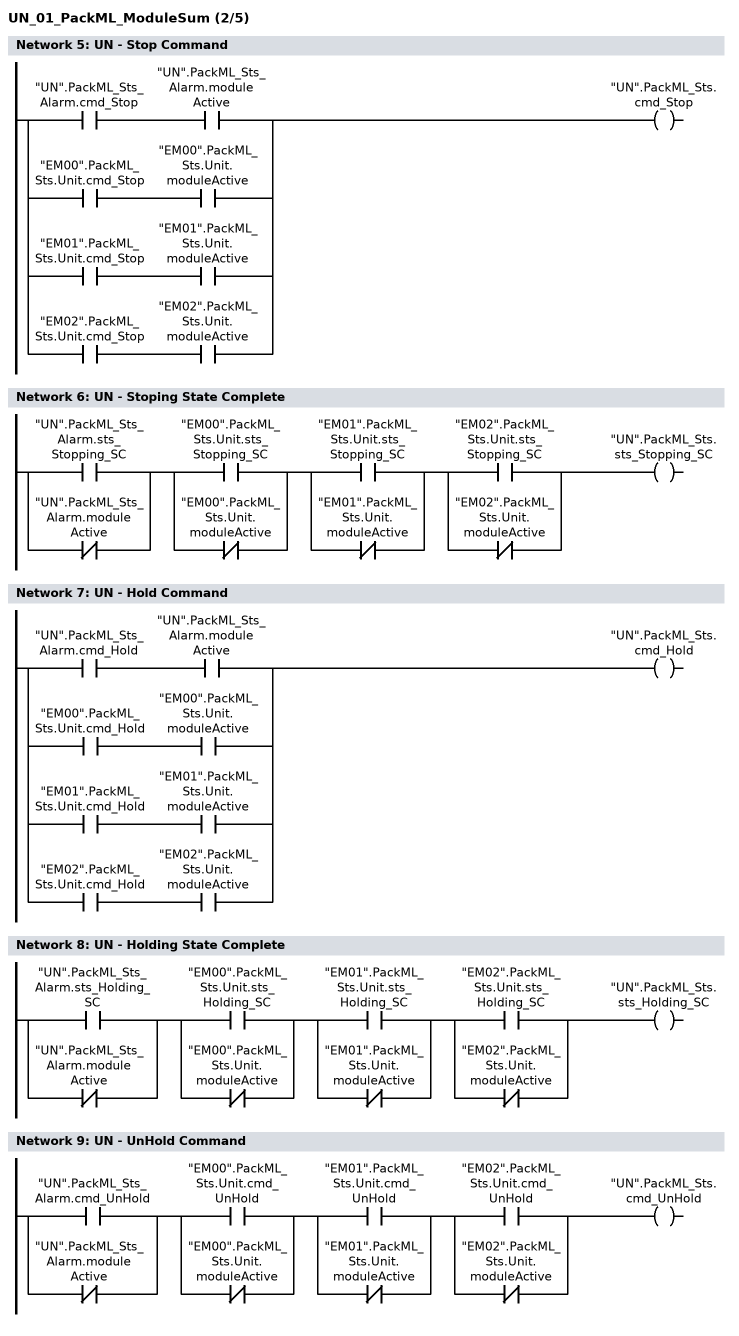
   RUNG wire#powerrail
      Contact( "UN".PackML_Sts_Alarm.cmd_Stop )
      Contact( "UN".PackML_Sts_Alarm.moduleActive )
      wire#w1
      Coil( "UN".PackML_Sts.cmd_Stop )
   END_RUNG
   RUNG wire#powerrail
      Contact( "EM00".PackML_Sts.Unit.cmd_Stop )
      Contact( "EM00".PackML_Sts.Unit.moduleActive )
   END_RUNG wire#w1
   RUNG wire#powerrail
      Contact( "EM01".PackML_Sts.Unit.cmd_Stop )
      Contact( "EM01".PackML_Sts.Unit.moduleActive )
   END_RUNG wire#w1
   RUNG wire#powerrail
      Contact( "EM02".PackML_Sts.Unit.cmd_Stop )
      Contact( "EM02".PackML_Sts.Unit.moduleActive )
   END_RUNG wire#w1
   // the same network as SCL:
   "UN".PackML_Sts.cmd_Stop := ("UN".PackML_Sts_Alarm.cmd_Stop AND "UN".PackML_Sts_Alarm.moduleActive) OR ("EM00".PackML_Sts.Unit.cmd_Stop AND "EM00".PackML_Sts.Unit.moduleActive) OR ("EM01".PackML_Sts.Unit.cmd_Stop AND "EM01".PackML_Sts.Unit.moduleActive) OR ("EM02".PackML_Sts.Unit.cmd_Stop AND "EM02".PackML_Sts.Unit.moduleActive);
END_REGION

REGION Network 6: UN - Stoping State Complete
   RUNG wire#powerrail
      Contact( "UN".PackML_Sts_Alarm.sts_Stopping_SC )
      wire#w1
      Contact( "EM00".PackML_Sts.Unit.sts_Stopping_SC )
      wire#w2
      Contact( "EM01".PackML_Sts.Unit.sts_Stopping_SC )
      wire#w3
      Contact( "EM02".PackML_Sts.Unit.sts_Stopping_SC )
      wire#w4
      Coil( "UN".PackML_Sts.sts_Stopping_SC )
   END_RUNG
   RUNG wire#powerrail
      I_Contact( "UN".PackML_Sts_Alarm.moduleActive )
   END_RUNG wire#w1
   RUNG wire#w1
      I_Contact( "EM00".PackML_Sts.Unit.moduleActive )
   END_RUNG wire#w2
   RUNG wire#w2
      I_Contact( "EM01".PackML_Sts.Unit.moduleActive )
   END_RUNG wire#w3
   RUNG wire#w3
      I_Contact( "EM02".PackML_Sts.Unit.moduleActive )
   END_RUNG wire#w4
   // the same network as SCL:
   "UN".PackML_Sts.sts_Stopping_SC := ("UN".PackML_Sts_Alarm.sts_Stopping_SC OR NOT "UN".PackML_Sts_Alarm.moduleActive) AND ("EM00".PackML_Sts.Unit.sts_Stopping_SC OR NOT "EM00".PackML_Sts.Unit.moduleActive) AND ("EM01".PackML_Sts.Unit.sts_Stopping_SC OR NOT "EM01".PackML_Sts.Unit.moduleActive) AND ("EM02".PackML_Sts.Unit.sts_Stopping_SC OR NOT "EM02".PackML_Sts.Unit.moduleActive);
END_REGION
